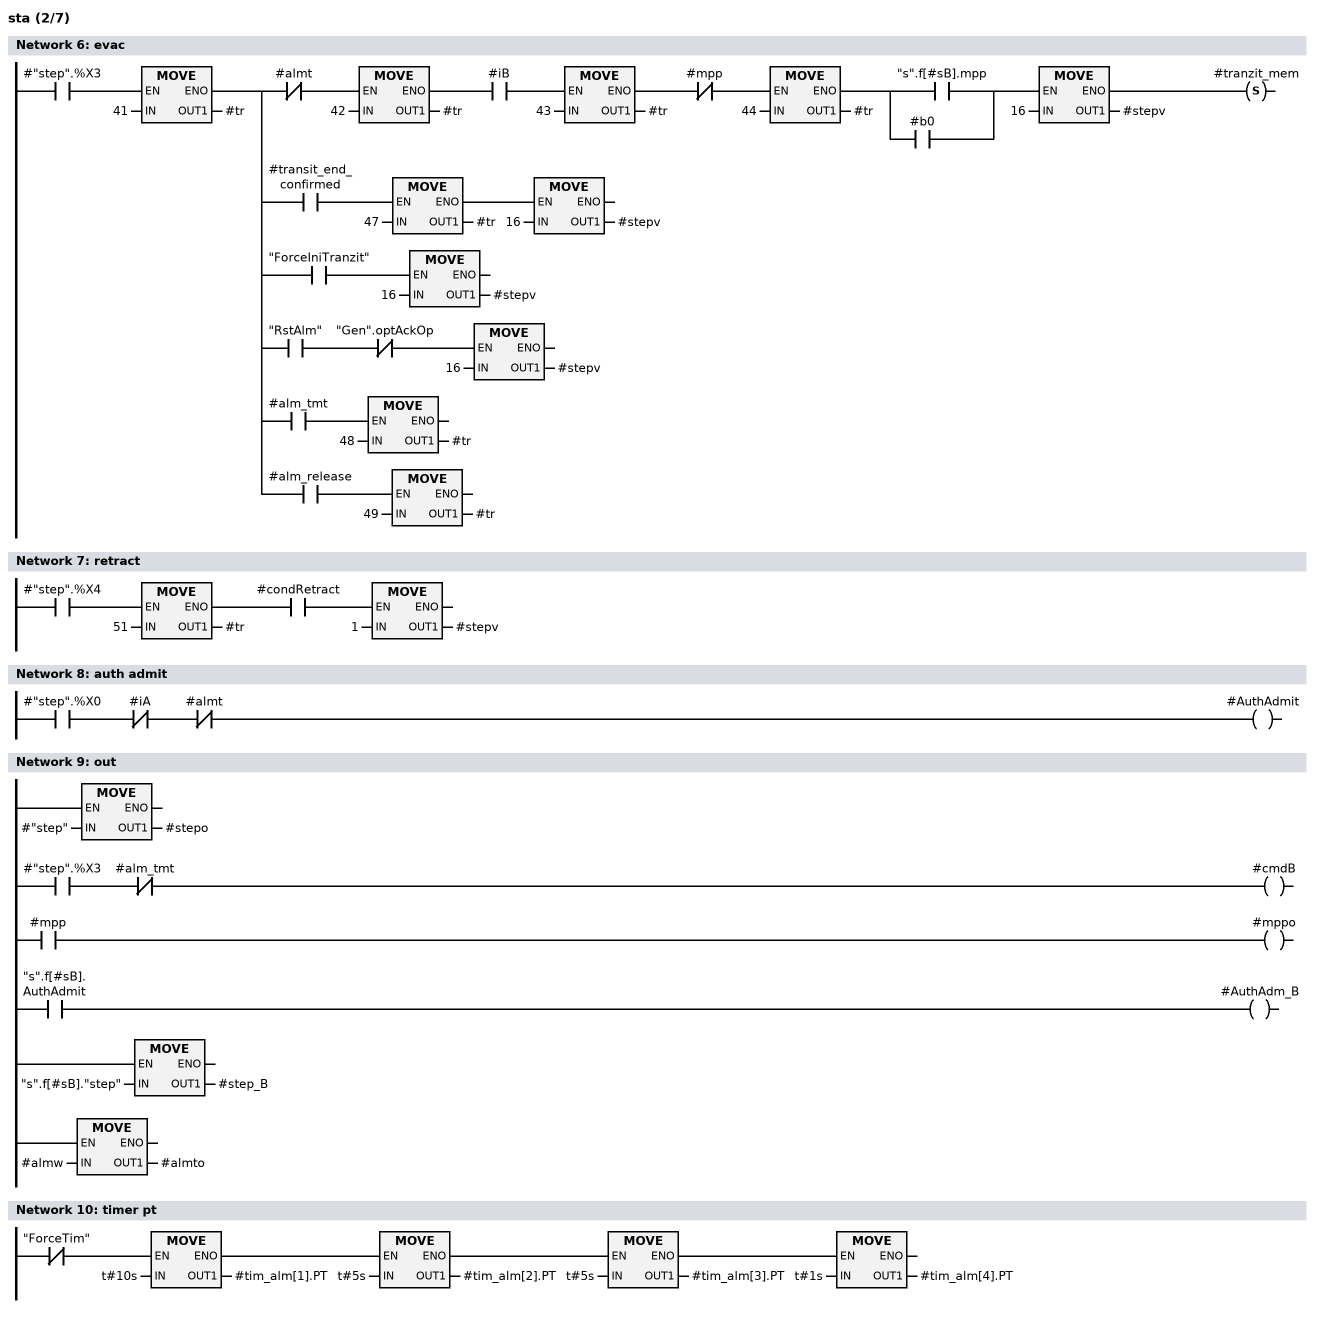
   RUNG wire#powerrail
      Contact( #"step".%X3 )
      Move(in := 41, out1 => #tr)
      wire#w1
      I_Contact( #almt )
      Move(in := 42, out1 => #tr)
      Contact( #iB )
      Move(in := 43, out1 => #tr)
      I_Contact( #mpp )
      Move(in := 44, out1 => #tr)
      wire#w2
      Contact( "s".f[#sB].mpp )
      wire#w3
      Move(in := 16, out1 => #stepv)
      S_Coil( #tranzit_mem )
   END_RUNG
   RUNG wire#w2
      Contact( #b0 )
   END_RUNG wire#w3
   RUNG wire#w1
      Contact( #transit_end_confirmed )
      Move(in := 47, out1 => #tr)
      Move(in := 16, out1 => #stepv)
   END_RUNG
   RUNG wire#w1
      Contact( "ForceIniTranzit" )
      Move(in := 16, out1 => #stepv)
   END_RUNG
   RUNG wire#w1
      Contact( "RstAlm" )
      I_Contact( "Gen".optAckOp )
      Move(in := 16, out1 => #stepv)
   END_RUNG
   RUNG wire#w1
      Contact( #alm_tmt )
      Move(in := 48, out1 => #tr)
   END_RUNG
   RUNG wire#w1
      Contact( #alm_release )
      Move(in := 49, out1 => #tr)
   END_RUNG
   // the same network as SCL:
   IF #"step".%X3 THEN #tr := 41; END_IF;
   #_w1 := #"step".%X3 AND NOT #almt;
   IF #_w1 THEN #tr := 42; END_IF;
   #_w2 := #_w1 AND #iB;
   IF #_w2 THEN #tr := 43; END_IF;
   #_w3 := #_w2 AND NOT #mpp;
   IF #_w3 THEN #tr := 44; END_IF;
   IF #_w3 AND ("s".f[#sB].mpp OR #b0) THEN
       #stepv := 16;
       #tranzit_mem := TRUE;
   END_IF;
   IF #"step".%X3 AND #transit_end_confirmed THEN
       #tr := 47;
       #stepv := 16;
   END_IF;
   IF #"step".%X3 AND "ForceIniTranzit" THEN #stepv := 16; END_IF;
   IF #"step".%X3 AND "RstAlm" AND NOT "Gen".optAckOp THEN #stepv := 16; END_IF;
   IF #"step".%X3 AND #alm_tmt THEN #tr := 48; END_IF;
   IF #"step".%X3 AND #alm_release THEN #tr := 49; END_IF;
END_REGION

REGION Network 7: retract
   RUNG wire#powerrail
      Contact( #"step".%X4 )
      Move(in := 51, out1 => #tr)
      Contact( #condRetract )
      Move(in := 1, out1 => #stepv)
   END_RUNG
   // the same network as SCL:
   IF #"step".%X4 THEN #tr := 51; END_IF;
   IF #"step".%X4 AND #condRetract THEN #stepv := 1; END_IF;
END_REGION

REGION Network 8: auth admit
   RUNG wire#powerrail
      Contact( #"step".%X0 )
      I_Contact( #iA )
      I_Contact( #almt )
      Coil( #AuthAdmit )
   END_RUNG
   // the same network as SCL:
   #AuthAdmit := #"step".%X0 AND NOT #iA AND NOT #almt;
END_REGION

REGION Network 9: out
   RUNG wire#powerrail
      Move(in := #"step", out1 => #stepo)
   END_RUNG
   RUNG wire#powerrail
      Contact( #"step".%X3 )
      I_Contact( #alm_tmt )
      Coil( #cmdB )
   END_RUNG
   RUNG wire#powerrail
      Contact( #mpp )
      Coil( #mppo )
   END_RUNG
   RUNG wire#powerrail
      Contact( "s".f[#sB].AuthAdmit )
      Coil( #AuthAdm_B )
   END_RUNG
   RUNG wire#powerrail
      Move(in := "s".f[#sB]."step", out1 => #step_B)
   END_RUNG
   RUNG wire#powerrail
      Move(in := #almw, out1 => #almto)
   END_RUNG
   // the same network as SCL:
   #stepo := #"step";
   #cmdB := #"step".%X3 AND NOT #alm_tmt;
   #mppo := #mpp;
   #AuthAdm_B := "s".f[#sB].AuthAdmit;
   #step_B := "s".f[#sB]."step";
   #almto := #almw;
END_REGION

REGION Network 10: timer pt
   RUNG wire#powerrail
      I_Contact( "ForceTim" )
      Move(in := t#10s, out1 => #tim_alm[1].PT)
      Move(in := t#5s, out1 => #tim_alm[2].PT)
      Move(in := t#5s, out1 => #tim_alm[3].PT)
      Move(in := t#1s, out1 => #tim_alm[4].PT)
   END_RUNG
   // the same network as SCL:
   IF NOT "ForceTim" THEN
       #tim_alm[1].PT := t#10s;
       #tim_alm[2].PT := t#5s;
       #tim_alm[3].PT := t#5s;
       #tim_alm[4].PT := t#1s;
   END_IF;
END_REGION

REGION Network 11: rst all
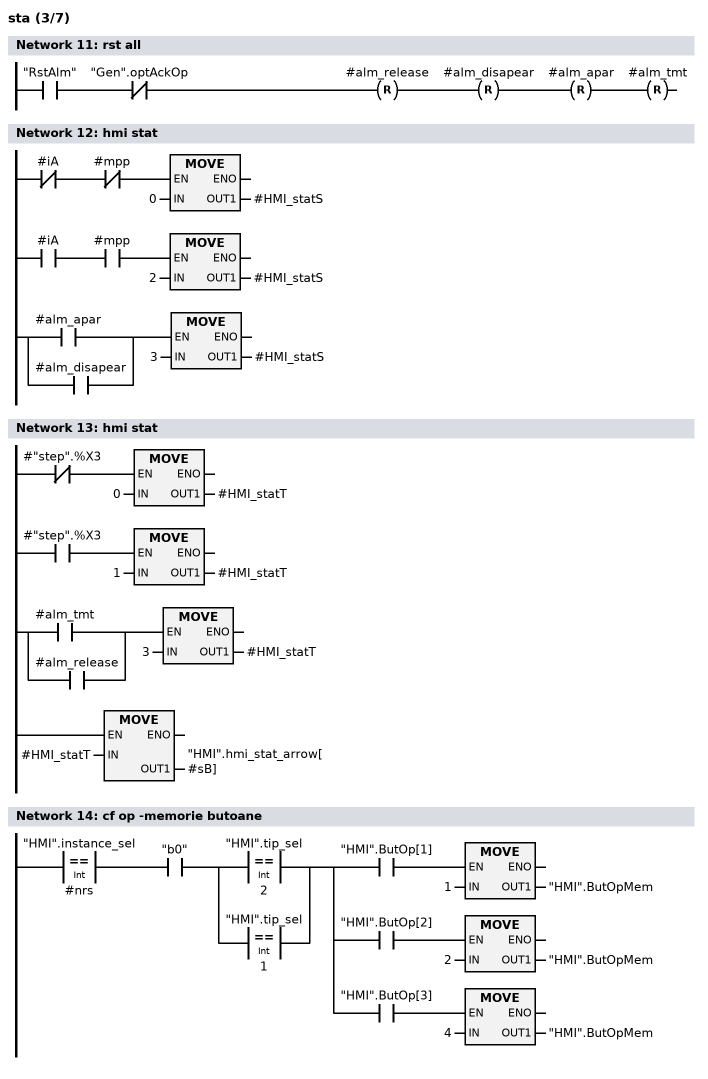
   RUNG wire#powerrail
      Contact( "RstAlm" )
      I_Contact( "Gen".optAckOp )
      R_Coil( #alm_release )
      R_Coil( #alm_disapear )
      R_Coil( #alm_apar )
      R_Coil( #alm_tmt )
   END_RUNG
   // the same network as SCL:
   IF "RstAlm" AND NOT "Gen".optAckOp THEN
       #alm_release := FALSE;
       #alm_disapear := FALSE;
       #alm_apar := FALSE;
       #alm_tmt := FALSE;
   END_IF;
END_REGION

REGION Network 12: hmi stat
   RUNG wire#powerrail
      I_Contact( #iA )
      I_Contact( #mpp )
      Move(in := 0, out1 => #HMI_statS)
   END_RUNG
   RUNG wire#powerrail
      Contact( #iA )
      Contact( #mpp )
      Move(in := 2, out1 => #HMI_statS)
   END_RUNG
   RUNG wire#powerrail
      Contact( #alm_apar )
      wire#w1
      Move(in := 3, out1 => #HMI_statS)
   END_RUNG
   RUNG wire#powerrail
      Contact( #alm_disapear )
   END_RUNG wire#w1
   // the same network as SCL:
   IF NOT #iA AND NOT #mpp THEN #HMI_statS := 0; END_IF;
   IF #iA AND #mpp THEN #HMI_statS := 2; END_IF;
   IF #alm_apar OR #alm_disapear THEN #HMI_statS := 3; END_IF;
END_REGION

REGION Network 13: hmi stat
   RUNG wire#powerrail
      I_Contact( #"step".%X3 )
      Move(in := 0, out1 => #HMI_statT)
   END_RUNG
   RUNG wire#powerrail
      Contact( #"step".%X3 )
      Move(in := 1, out1 => #HMI_statT)
   END_RUNG
   RUNG wire#powerrail
      Contact( #alm_tmt )
      wire#w1
      Move(in := 3, out1 => #HMI_statT)
   END_RUNG
   RUNG wire#powerrail
      Contact( #alm_release )
   END_RUNG wire#w1
   RUNG wire#powerrail
      Move(in := #HMI_statT, out1 => "HMI".hmi_stat_arrow[#sB])
   END_RUNG
   // the same network as SCL:
   IF NOT #"step".%X3 THEN #HMI_statT := 0; END_IF;
   IF #"step".%X3 THEN #HMI_statT := 1; END_IF;
   IF #alm_tmt OR #alm_release THEN #HMI_statT := 3; END_IF;
   "HMI".hmi_stat_arrow[#sB] := #HMI_statT;
END_REGION

REGION Network 14: cf op -memorie butoane
   RUNG wire#powerrail
      { S7_Templates := "SrcType := Int" } EQ_Contact(in1 := "HMI".instance_sel, in2 := #nrs)
      Contact( "b0" )
      wire#w1
      { S7_Templates := "SrcType := Int" } EQ_Contact(in1 := "HMI".tip_sel, in2 := 2)
      wire#w2
      Contact( "HMI".ButOp[1] )
      Move(in := 1, out1 => "HMI".ButOpMem)
   END_RUNG
   RUNG wire#w1
      { S7_Templates := "SrcType := Int" } EQ_Contact(in1 := "HMI".tip_sel, in2 := 1)
   END_RUNG wire#w2
   RUNG wire#w2
      Contact( "HMI".ButOp[2] )
      Move(in := 2, out1 => "HMI".ButOpMem)
   END_RUNG
   RUNG wire#w2
      Contact( "HMI".ButOp[3] )
      Move(in := 4, out1 => "HMI".ButOpMem)
   END_RUNG
   // the same network as SCL:
   #_w1 := ("HMI".instance_sel = #nrs) AND "b0" AND (("HMI".tip_sel = 2) OR ("HMI".tip_sel = 1));
   IF #_w1 AND "HMI".ButOp[1] THEN "HMI".ButOpMem := 1; END_IF;
   IF #_w1 AND "HMI".ButOp[2] THEN "HMI".ButOpMem := 2; END_IF;
   IF #_w1 AND "HMI".ButOp[3] THEN "HMI".ButOpMem := 4; END_IF;
END_REGION

REGION Network 15: cf op alm tmt / release
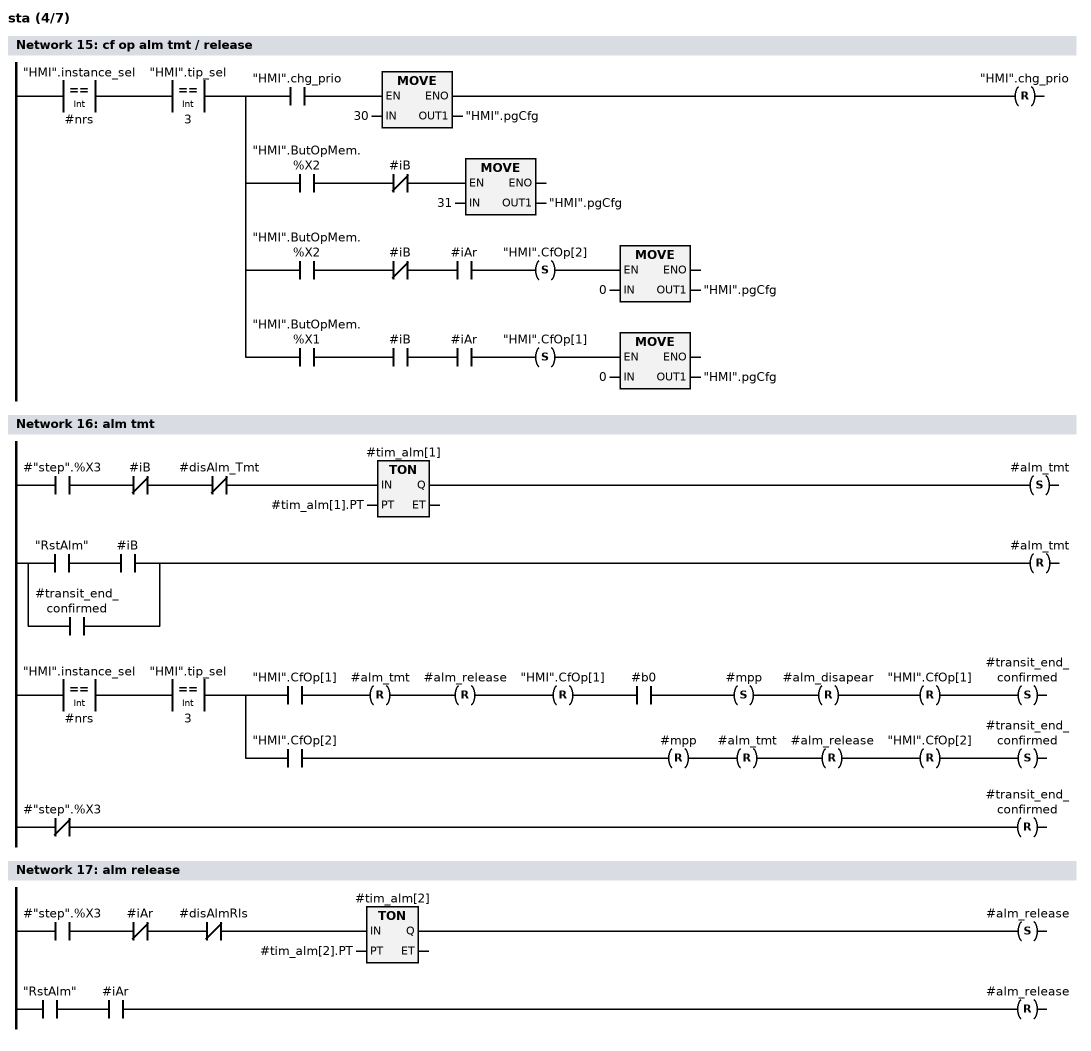
   RUNG wire#powerrail
      { S7_Templates := "SrcType := Int" } EQ_Contact(in1 := "HMI".instance_sel, in2 := #nrs)
      { S7_Templates := "SrcType := Int" } EQ_Contact(in1 := "HMI".tip_sel, in2 := 3)
      wire#w1
      Contact( "HMI".chg_prio )
      Move(in := 30, out1 => "HMI".pgCfg)
      R_Coil( "HMI".chg_prio )
   END_RUNG
   RUNG wire#w1
      Contact( "HMI".ButOpMem.%X2 )
      I_Contact( #iB )
      Move(in := 31, out1 => "HMI".pgCfg)
   END_RUNG
   RUNG wire#w1
      Contact( "HMI".ButOpMem.%X2 )
      I_Contact( #iB )
      Contact( #iAr )
      S_Coil( "HMI".CfOp[2] )
      Move(in := 0, out1 => "HMI".pgCfg)
   END_RUNG
   RUNG wire#w1
      Contact( "HMI".ButOpMem.%X1 )
      Contact( #iB )
      Contact( #iAr )
      S_Coil( "HMI".CfOp[1] )
      Move(in := 0, out1 => "HMI".pgCfg)
   END_RUNG
   // the same network as SCL:
   #_w1 := ("HMI".instance_sel = #nrs) AND ("HMI".tip_sel = 3);
   IF #_w1 AND "HMI".chg_prio THEN
       "HMI".pgCfg := 30;
       "HMI".chg_prio := FALSE;
   END_IF;
   IF #_w1 AND "HMI".ButOpMem.%X2 AND NOT #iB THEN "HMI".pgCfg := 31; END_IF;
   IF #_w1 AND "HMI".ButOpMem.%X2 AND NOT #iB AND #iAr THEN
       "HMI".CfOp[2] := TRUE;
       "HMI".pgCfg := 0;
   END_IF;
   IF #_w1 AND "HMI".ButOpMem.%X1 AND #iB AND #iAr THEN
       "HMI".CfOp[1] := TRUE;
       "HMI".pgCfg := 0;
   END_IF;
END_REGION

REGION Network 16: alm tmt
   #tim_alm[1].TON(IN := #"step".%X3 AND NOT #iB AND NOT #disAlm_Tmt, PT := #tim_alm[1].PT);
   IF #tim_alm[1].Q THEN #alm_tmt := TRUE; END_IF;
   IF ("RstAlm" AND #iB) OR #transit_end_confirmed THEN #alm_tmt := FALSE; END_IF;
   #_w1 := ("HMI".instance_sel = #nrs) AND ("HMI".tip_sel = 3);
   #_w2 := #_w1 AND "HMI".CfOp[1];
   IF #_w2 THEN
       #alm_tmt := FALSE;
       #alm_release := FALSE;
       "HMI".CfOp[1] := FALSE;
   END_IF;
   IF #_w2 AND #b0 THEN
       #mpp := TRUE;
       #alm_disapear := FALSE;
       "HMI".CfOp[1] := FALSE;
       #transit_end_confirmed := TRUE;
   END_IF;
   IF #_w1 AND "HMI".CfOp[2] THEN
       #mpp := FALSE;
       #alm_tmt := FALSE;
       #alm_release := FALSE;
   END_IF;
   #_w3 := #_w1 AND "HMI".CfOp[2];
   IF #_w3 THEN
       "HMI".CfOp[2] := FALSE;
       #transit_end_confirmed := TRUE;
   END_IF;
   IF NOT #"step".%X3 THEN #transit_end_confirmed := FALSE; END_IF;
END_REGION

REGION Network 17: alm release
   #tim_alm[2].TON(IN := #"step".%X3 AND NOT #iAr AND NOT #disAlmRls, PT := #tim_alm[2].PT);
   IF #tim_alm[2].Q THEN #alm_release := TRUE; END_IF;
   IF "RstAlm" AND #iAr THEN #alm_release := FALSE; END_IF;
END_REGION

REGION Network 18: cf op alarma disparitie fara tranzit
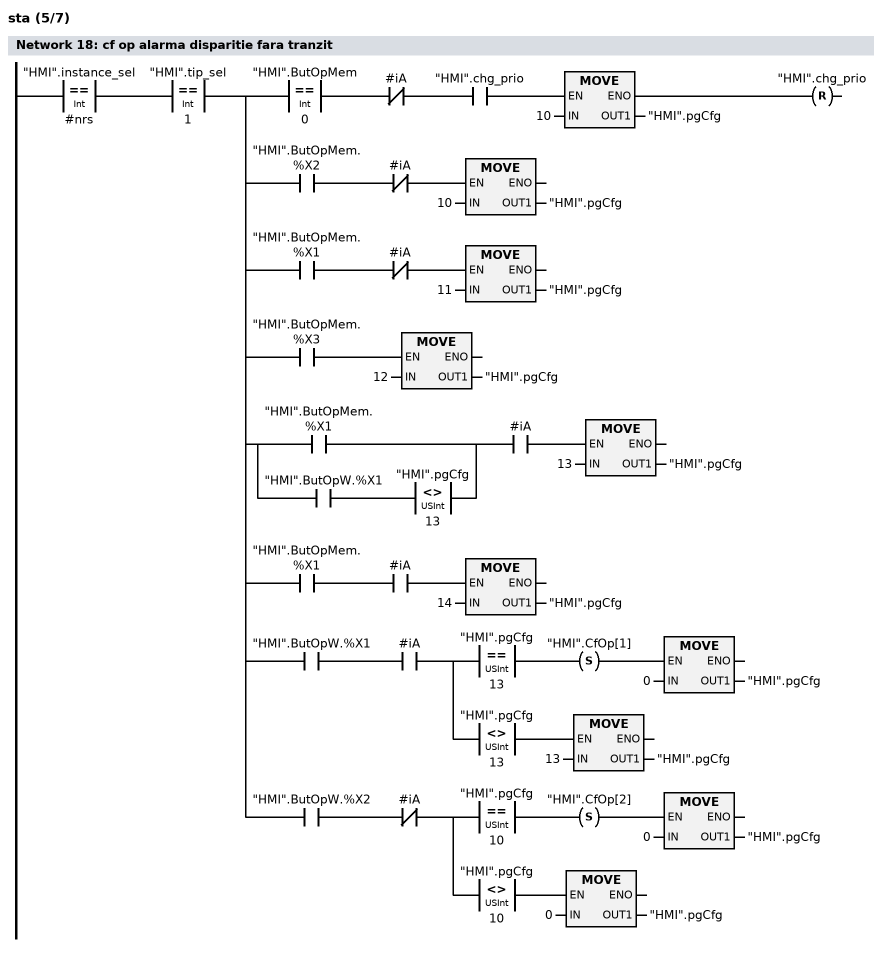
   RUNG wire#powerrail
      { S7_Templates := "SrcType := Int" } EQ_Contact(in1 := "HMI".instance_sel, in2 := #nrs)
      { S7_Templates := "SrcType := Int" } EQ_Contact(in1 := "HMI".tip_sel, in2 := 1)
      wire#w1
      { S7_Templates := "SrcType := Int" } EQ_Contact(in1 := "HMI".ButOpMem, in2 := 0)
      I_Contact( #iA )
      Contact( "HMI".chg_prio )
      Move(in := 10, out1 => "HMI".pgCfg)
      R_Coil( "HMI".chg_prio )
   END_RUNG
   RUNG wire#w1
      Contact( "HMI".ButOpMem.%X2 )
      I_Contact( #iA )
      Move(in := 10, out1 => "HMI".pgCfg)
   END_RUNG
   RUNG wire#w1
      Contact( "HMI".ButOpMem.%X1 )
      I_Contact( #iA )
      Move(in := 11, out1 => "HMI".pgCfg)
   END_RUNG
   RUNG wire#w1
      Contact( "HMI".ButOpMem.%X3 )
      Move(in := 12, out1 => "HMI".pgCfg)
   END_RUNG
   RUNG wire#w1
      Contact( "HMI".ButOpMem.%X1 )
      wire#w2
      Contact( #iA )
      Move(in := 13, out1 => "HMI".pgCfg)
   END_RUNG
   RUNG wire#w1
      Contact( "HMI".ButOpW.%X1 )
      { S7_Templates := "SrcType := USInt" } NE_Contact(in1 := "HMI".pgCfg, in2 := 13)
   END_RUNG wire#w2
   RUNG wire#w1
      Contact( "HMI".ButOpMem.%X1 )
      Contact( #iA )
      Move(in := 14, out1 => "HMI".pgCfg)
   END_RUNG
   RUNG wire#w1
      Contact( "HMI".ButOpW.%X1 )
      Contact( #iA )
      wire#w3
      { S7_Templates := "SrcType := USInt" } EQ_Contact(in1 := "HMI".pgCfg, in2 := 13)
      S_Coil( "HMI".CfOp[1] )
      Move(in := 0, out1 => "HMI".pgCfg)
   END_RUNG
   RUNG wire#w3
      { S7_Templates := "SrcType := USInt" } NE_Contact(in1 := "HMI".pgCfg, in2 := 13)
      Move(in := 13, out1 => "HMI".pgCfg)
   END_RUNG
   RUNG wire#w1
      Contact( "HMI".ButOpW.%X2 )
      I_Contact( #iA )
      wire#w4
      { S7_Templates := "SrcType := USInt" } EQ_Contact(in1 := "HMI".pgCfg, in2 := 10)
      S_Coil( "HMI".CfOp[2] )
      Move(in := 0, out1 => "HMI".pgCfg)
   END_RUNG
   RUNG wire#w4
      { S7_Templates := "SrcType := USInt" } NE_Contact(in1 := "HMI".pgCfg, in2 := 10)
      Move(in := 0, out1 => "HMI".pgCfg)
   END_RUNG
   // the same network as SCL:
   #_w1 := ("HMI".instance_sel = #nrs) AND ("HMI".tip_sel = 1);
   IF #_w1 AND ("HMI".ButOpMem = 0) AND NOT #iA AND "HMI".chg_prio THEN
       "HMI".pgCfg := 10;
       "HMI".chg_prio := FALSE;
   END_IF;
   IF #_w1 AND "HMI".ButOpMem.%X2 AND NOT #iA THEN "HMI".pgCfg := 10; END_IF;
   IF #_w1 AND "HMI".ButOpMem.%X1 AND NOT #iA THEN "HMI".pgCfg := 11; END_IF;
   IF #_w1 AND "HMI".ButOpMem.%X3 THEN "HMI".pgCfg := 12; END_IF;
   IF #_w1 AND ("HMI".ButOpMem.%X1 OR ("HMI".ButOpW.%X1 AND ("HMI".pgCfg <> 13))) AND #iA THEN
       "HMI".pgCfg := 13;
   END_IF;
   IF #_w1 AND "HMI".ButOpMem.%X1 AND #iA THEN "HMI".pgCfg := 14; END_IF;
   #_w2 := #_w1 AND "HMI".ButOpW.%X1 AND #iA;
   IF #_w2 AND ("HMI".pgCfg = 13) THEN
       "HMI".CfOp[1] := TRUE;
       "HMI".pgCfg := 0;
   END_IF;
   IF #_w2 AND ("HMI".pgCfg <> 13) THEN "HMI".pgCfg := 13; END_IF;
   #_w3 := #_w1 AND "HMI".ButOpW.%X2 AND NOT #iA;
   IF #_w3 AND ("HMI".pgCfg = 10) THEN
       "HMI".CfOp[2] := TRUE;
       "HMI".pgCfg := 0;
   END_IF;
   IF #_w3 AND ("HMI".pgCfg <> 10) THEN "HMI".pgCfg := 0; END_IF;
END_REGION

REGION Network 19: alm disap
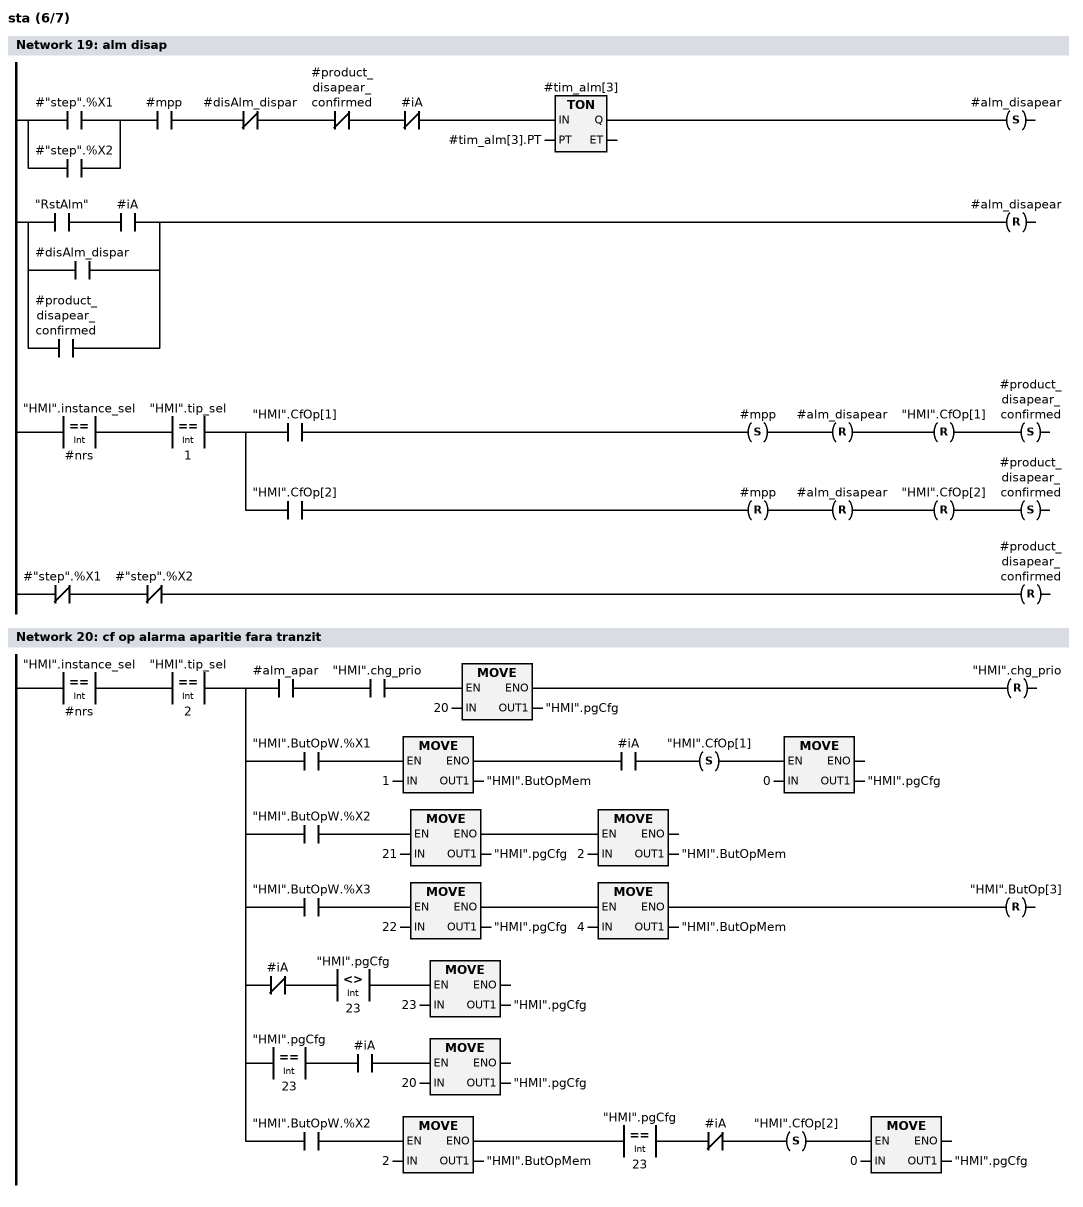
   #tim_alm[3].TON(IN := (#"step".%X1 OR #"step".%X2) AND #mpp AND NOT #disAlm_dispar AND NOT #product_disapear_confirmed AND NOT #iA,
                   PT := #tim_alm[3].PT);
   IF #tim_alm[3].Q THEN #alm_disapear := TRUE; END_IF;
   IF ("RstAlm" AND #iA) OR #disAlm_dispar OR #product_disapear_confirmed THEN
       #alm_disapear := FALSE;
   END_IF;
   #_w1 := ("HMI".instance_sel = #nrs) AND ("HMI".tip_sel = 1);
   IF #_w1 AND "HMI".CfOp[1] THEN
       #mpp := TRUE;
       #alm_disapear := FALSE;
   END_IF;
   #_w2 := #_w1 AND "HMI".CfOp[1];
   IF #_w2 THEN
       "HMI".CfOp[1] := FALSE;
       #product_disapear_confirmed := TRUE;
   END_IF;
   IF #_w1 AND "HMI".CfOp[2] THEN
       #mpp := FALSE;
       #alm_disapear := FALSE;
   END_IF;
   #_w3 := #_w1 AND "HMI".CfOp[2];
   IF #_w3 THEN
       "HMI".CfOp[2] := FALSE;
       #product_disapear_confirmed := TRUE;
   END_IF;
   IF NOT #"step".%X1 AND NOT #"step".%X2 THEN #product_disapear_confirmed := FALSE; END_IF;
END_REGION

REGION Network 20: cf op alarma aparitie fara tranzit
   RUNG wire#powerrail
      { S7_Templates := "SrcType := Int" } EQ_Contact(in1 := "HMI".instance_sel, in2 := #nrs)
      { S7_Templates := "SrcType := Int" } EQ_Contact(in1 := "HMI".tip_sel, in2 := 2)
      wire#w1
      Contact( #alm_apar )
      Contact( "HMI".chg_prio )
      Move(in := 20, out1 => "HMI".pgCfg)
      R_Coil( "HMI".chg_prio )
   END_RUNG
   RUNG wire#w1
      Contact( "HMI".ButOpW.%X1 )
      Move(in := 1, out1 => "HMI".ButOpMem)
      Contact( #iA )
      S_Coil( "HMI".CfOp[1] )
      Move(in := 0, out1 => "HMI".pgCfg)
   END_RUNG
   RUNG wire#w1
      Contact( "HMI".ButOpW.%X2 )
      Move(in := 21, out1 => "HMI".pgCfg)
      Move(in := 2, out1 => "HMI".ButOpMem)
   END_RUNG
   RUNG wire#w1
      Contact( "HMI".ButOpW.%X3 )
      Move(in := 22, out1 => "HMI".pgCfg)
      Move(in := 4, out1 => "HMI".ButOpMem)
      R_Coil( "HMI".ButOp[3] )
   END_RUNG
   RUNG wire#w1
      I_Contact( #iA )
      { S7_Templates := "SrcType := Int" } NE_Contact(in1 := "HMI".pgCfg, in2 := 23)
      Move(in := 23, out1 => "HMI".pgCfg)
   END_RUNG
   RUNG wire#w1
      { S7_Templates := "SrcType := Int" } EQ_Contact(in1 := "HMI".pgCfg, in2 := 23)
      Contact( #iA )
      Move(in := 20, out1 => "HMI".pgCfg)
   END_RUNG
   RUNG wire#w1
      Contact( "HMI".ButOpW.%X2 )
      Move(in := 2, out1 => "HMI".ButOpMem)
      { S7_Templates := "SrcType := Int" } EQ_Contact(in1 := "HMI".pgCfg, in2 := 23)
      I_Contact( #iA )
      S_Coil( "HMI".CfOp[2] )
      Move(in := 0, out1 => "HMI".pgCfg)
   END_RUNG
   // the same network as SCL:
   #_w1 := ("HMI".instance_sel = #nrs) AND ("HMI".tip_sel = 2);
   IF #_w1 AND #alm_apar AND "HMI".chg_prio THEN
       "HMI".pgCfg := 20;
       "HMI".chg_prio := FALSE;
   END_IF;
   #_w2 := #_w1 AND "HMI".ButOpW.%X1;
   IF #_w2 THEN "HMI".ButOpMem := 1; END_IF;
   IF #_w2 AND #iA THEN
       "HMI".CfOp[1] := TRUE;
       "HMI".pgCfg := 0;
   END_IF;
   IF #_w1 AND "HMI".ButOpW.%X2 THEN
       "HMI".pgCfg := 21;
       "HMI".ButOpMem := 2;
   END_IF;
   IF #_w1 AND "HMI".ButOpW.%X3 THEN
       "HMI".pgCfg := 22;
       "HMI".ButOpMem := 4;
       "HMI".ButOp[3] := FALSE;
   END_IF;
   IF #_w1 AND NOT #iA AND ("HMI".pgCfg <> 23) THEN "HMI".pgCfg := 23; END_IF;
   IF #_w1 AND ("HMI".pgCfg = 23) AND #iA THEN "HMI".pgCfg := 20; END_IF;
   #_w3 := #_w1 AND "HMI".ButOpW.%X2;
   IF #_w3 THEN "HMI".ButOpMem := 2; END_IF;
   IF #_w3 AND ("HMI".pgCfg = 23) AND NOT #iA THEN
       "HMI".CfOp[2] := TRUE;
       "HMI".pgCfg := 0;
   END_IF;
END_REGION

REGION Network 21: alm apar
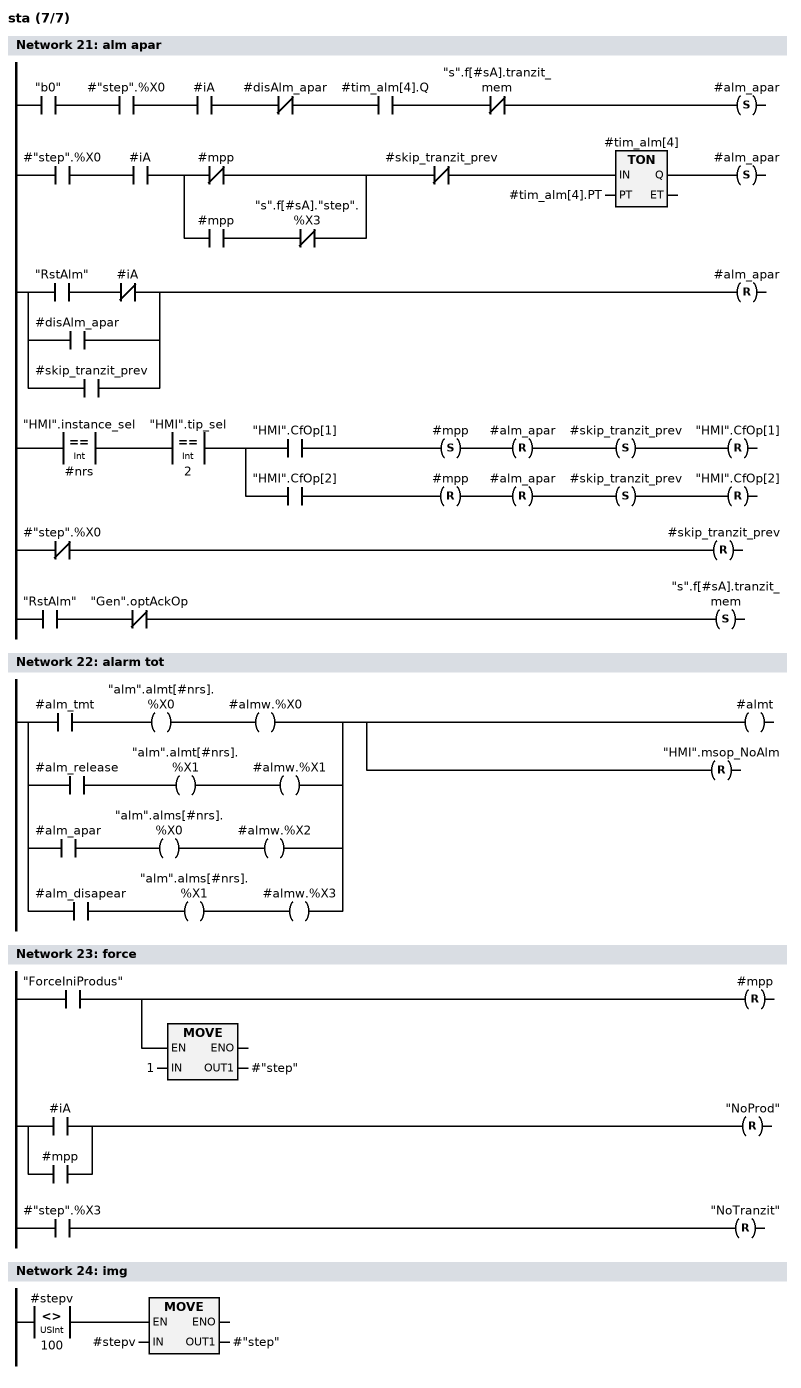
   IF "b0" AND #"step".%X0 AND #iA AND NOT #disAlm_apar AND #tim_alm[4].Q AND NOT "s".f[#sA].tranzit_mem THEN
       #alm_apar := TRUE;
   END_IF;
   #tim_alm[4].TON(IN := #"step".%X0 AND #iA AND (NOT #mpp OR (#mpp AND NOT "s".f[#sA]."step".%X3)) AND NOT #skip_tranzit_prev,
                   PT := #tim_alm[4].PT);
   IF #tim_alm[4].Q THEN #alm_apar := TRUE; END_IF;
   IF ("RstAlm" AND NOT #iA) OR #disAlm_apar OR #skip_tranzit_prev THEN #alm_apar := FALSE; END_IF;
   #_w1 := ("HMI".instance_sel = #nrs) AND ("HMI".tip_sel = 2);
   IF #_w1 AND "HMI".CfOp[1] THEN
       #mpp := TRUE;
       #alm_apar := FALSE;
       #skip_tranzit_prev := TRUE;
       "HMI".CfOp[1] := FALSE;
   END_IF;
   IF #_w1 AND "HMI".CfOp[2] THEN
       #mpp := FALSE;
       #alm_apar := FALSE;
       #skip_tranzit_prev := TRUE;
       "HMI".CfOp[2] := FALSE;
   END_IF;
   IF NOT #"step".%X0 THEN #skip_tranzit_prev := FALSE; END_IF;
   IF "RstAlm" AND NOT "Gen".optAckOp THEN "s".f[#sA].tranzit_mem := TRUE; END_IF;
END_REGION

REGION Network 22: alarm tot
   RUNG wire#powerrail
      Contact( #alm_tmt )
      Coil( "alm".almt[#nrs].%X0 )
      Coil( #almw.%X0 )
      wire#w1
      Coil( #almt )
   END_RUNG
   RUNG wire#powerrail
      Contact( #alm_release )
      Coil( "alm".almt[#nrs].%X1 )
      Coil( #almw.%X1 )
   END_RUNG wire#w1
   RUNG wire#powerrail
      Contact( #alm_apar )
      Coil( "alm".alms[#nrs].%X0 )
      Coil( #almw.%X2 )
   END_RUNG wire#w1
   RUNG wire#powerrail
      Contact( #alm_disapear )
      Coil( "alm".alms[#nrs].%X1 )
      Coil( #almw.%X3 )
   END_RUNG wire#w1
   RUNG wire#w1
      R_Coil( "HMI".msop_NoAlm )
   END_RUNG
   // the same network as SCL:
   "alm".almt[#nrs].%X0 := #alm_tmt;
   #almw.%X0 := #alm_tmt;
   "alm".almt[#nrs].%X1 := #alm_release;
   #almw.%X1 := #alm_release;
   "alm".alms[#nrs].%X0 := #alm_apar;
   #almw.%X2 := #alm_apar;
   "alm".alms[#nrs].%X1 := #alm_disapear;
   #almw.%X3 := #alm_disapear;
   #almt := #alm_tmt OR #alm_release OR #alm_apar OR #alm_disapear;
   IF #almt THEN "HMI".msop_NoAlm := FALSE; END_IF;
END_REGION

REGION Network 23: force
   RUNG wire#powerrail
      Contact( "ForceIniProdus" )
      wire#w1
      R_Coil( #mpp )
   END_RUNG
   RUNG wire#w1
      Move(in := 1, out1 => #"step")
   END_RUNG
   RUNG wire#powerrail
      Contact( #iA )
      wire#w2
      R_Coil( "NoProd" )
   END_RUNG
   RUNG wire#powerrail
      Contact( #mpp )
   END_RUNG wire#w2
   RUNG wire#powerrail
      Contact( #"step".%X3 )
      R_Coil( "NoTranzit" )
   END_RUNG
   // the same network as SCL:
   IF "ForceIniProdus" THEN
       #mpp := FALSE;
       #"step" := 1;
   END_IF;
   IF #iA OR #mpp THEN "NoProd" := FALSE; END_IF;
   IF #"step".%X3 THEN "NoTranzit" := FALSE; END_IF;
END_REGION

REGION Network 24: img
   RUNG wire#powerrail
      { S7_Templates := "SrcType := USInt" } NE_Contact(in1 := #stepv, in2 := 100)
      Move(in := #stepv, out1 => #"step")
   END_RUNG
   // the same network as SCL:
   IF #stepv <> 100 THEN #"step" := #stepv; END_IF;
END_REGION
END_FUNCTION_BLOCK

FUNCTION_BLOCK "FB_GEN"   // FB14, LAD
{ S7_Optimized_Access := 'TRUE' }
VERSION : 0.1
   VAR
      tim : Array[1..15] of IEC_TIMER;
   END_VAR
   VAR_TEMP   // added for the SCL form of the ladder/FBD networks
      _w1 : Bool;
   END_VAR
BEGIN

REGION Network 1: Energie -Aer Z2_A
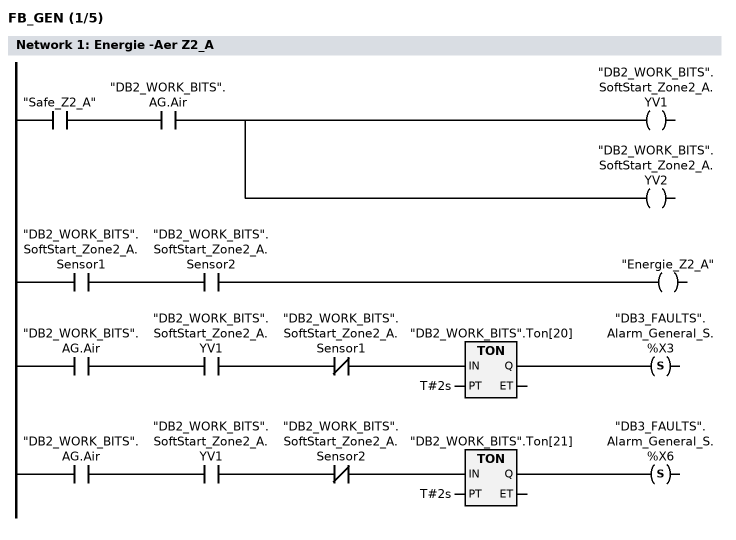
   "DB2_WORK_BITS".SoftStart_Zone2_A.YV1 := "Safe_Z2_A" AND "DB2_WORK_BITS".AG.Air;
   "DB2_WORK_BITS".SoftStart_Zone2_A.YV2 := "DB2_WORK_BITS".SoftStart_Zone2_A.YV1;
   "Energie_Z2_A" := "DB2_WORK_BITS".SoftStart_Zone2_A.Sensor1 AND "DB2_WORK_BITS".SoftStart_Zone2_A.Sensor2;
   "DB2_WORK_BITS".Ton[20].TON(IN := "DB2_WORK_BITS".AG.Air AND "DB2_WORK_BITS".SoftStart_Zone2_A.YV1 AND NOT "DB2_WORK_BITS".SoftStart_Zone2_A.Sensor1,
                           PT := T#2s);
   IF "DB2_WORK_BITS".Ton[20].Q THEN "DB3_FAULTS".Alarm_General_S.%X3 := TRUE; END_IF;
   "DB2_WORK_BITS".Ton[21].TON(IN := "DB2_WORK_BITS".AG.Air AND "DB2_WORK_BITS".SoftStart_Zone2_A.YV1 AND NOT "DB2_WORK_BITS".SoftStart_Zone2_A.Sensor2,
                           PT := T#2s);
   IF "DB2_WORK_BITS".Ton[21].Q THEN "DB3_FAULTS".Alarm_General_S.%X6 := TRUE; END_IF;
END_REGION

REGION Network 2: Energie -aer+power - Stack